TYPE "UDT1800_FLT_Machine"
VERSION : 0.1
   STRUCT
      Data_lost_after_erasing : Bool;   // Data_lost_after_erasing S7-CPU (1)
      Fuse_broken : Bool;   // Fuse broken machine (3)
      Connection_To_PC_lost : Bool;   // Connection to PC lost (3)
      Door_Swichtcabinet_open : Bool;   // Door swichtcabinet open(3)
      Air_dryer : Bool;   // Air dryer (3)
      Controlvoltage : Bool;   // Controlvoltage missing (M)
      CylinderServiceNotPermit : Bool;   // Operationmode cylinder service not permitted (1)
      Fuse_brocken_Mixinghead : Bool;   // Fuse broken mixinghead (3)
      Heating : Bool;   // Heating of machine overload (3)
      SGM_Faulty : Bool;   // Extrusion machine faulty (3)
      F_CoolingDevice : Bool;   // Compressor cooling device (3)
      WrongMH_No : Bool;   // Wrong mixinghead number (1)
      PlasmaFaulty : Bool;   // Plasma unit faulty (3)
      DrainingTank : Bool;   // Draining of a tank selected (M)
      SGM_AutomatcMissing : Bool;   // Extrusion machine not in automatic maode (3)
      Spare_1_7 : Bool;
      EmergencyStop : Struct   // Emergency stop general (M)
         Machine : Bool;   // Emergency stop nachine
         Switch_Cabinet : Bool;   // Emergency stop switch cabinet
         Operation_Panel : Bool;   // Emergency stop operation panel
         Monitor_2 : Bool;   // Emergency stop monitor_2
         Tank : Bool;   // Emergency stop tank
         MH_Cleaner_1 : Bool;   // Emergency stop mixinghead cleaner 1
         MH_Cleaner_2 : Bool;   // Emergency stop mixinghead cleaner 2
         Roboter_1 : Bool;   // Emergency stop Robot 1
         Roboter_2 : Bool;   // Emergency stop Robot 2
         ContStation_C1 : Bool;   // Emergency stop container station component 1
         ContStation_C2 : Bool;   // Emergency stop container station component 2
         External_Plant_1 : Bool;   // Emergency stop external plant 1
         External_Plant_2 : Bool;   // Emergency stop external plant 2
         ColorUnit_01 : Bool;   // Emergency stop color unit 1
         ColorUnit_02 : Bool;   // Emergency stop color unit 2
         AdditionalComponent : Bool;   // Emergency stop additional component
      END_STRUCT;
      OpMode_Test : Bool;   // Operation mode test is selected (M)
      Weekend_Mode : Bool;   // Weekende mode is active (M)
      Interface_PC : Bool;
      BufferBattery : Bool;
      AutoStop : Bool;   // AutoStop active (M)
      FLT_pre_alarm_pentan : Bool;   // Fault pre alarm pentan (3)
      FLT_alarm_pentan : Bool;   // Fault alarm pentan (1)
      P_AirSupply : Bool;   // Fault supply air pressure too low (3)
      FaultPC_Level_1 : Bool;
      FaultPC_Level_2 : Bool;
      FaultPC_Level_3 : Bool;
      Spare_13_3 : Bool;
      BufferShotDataFull : Bool;
      TransferFaultMMC : Bool;
      Fault_Watchdog : Bool;
      RefillStationNotReady : Bool;
      ShotTimeTooShort : Bool;
      CantDeleteTool : Bool;
      Pneumatik_1 : Bool;
      Pneumatik_2 : Bool;
      Spare_14_04 : Bool;
      Spare_14_05 : Bool;
      Spare_14_06 : Bool;
      Spare_14_07 : Bool;
      TimeValueIntervallNOK : Bool;
      Spare_15_01 : Bool;
      Spare_15_02 : Bool;
      Spare_15_03 : Bool;
      Spare_15_04 : Bool;
      Spare_15_05 : Bool;
      Spare_15_06 : Bool;
      Spare_15_07 : Bool;
      Spare_16_00 : Bool;
      Spare_16_01 : Bool;
      Spare_16_02 : Bool;
      Spare_16_03 : Bool;
      Spare_16_04 : Bool;
      Spare_16_05 : Bool;
      Spare_16_06 : Bool;
      Spare_16_07 : Bool;
      Spare_17_00 : Bool;
      Spare_17_01 : Bool;
      Spare_17_02 : Bool;
      Spare_17_03 : Bool;
      Spare_17_04 : Bool;
      Spare_17_05 : Bool;
      Spare_17_06 : Bool;
      Spare_17_07 : Bool;
   END_STRUCT;
END_TYPE

TYPE "UDT1801_FLT_auxDrive"
VERSION : 0.1
   STRUCT
      FLT_Motorprotection : Bool;   // Fault motorprotection
      FLT_FrequencyConverter : Bool;   // Fault frequency converter
      FLT_MaxP_MaxLTripTray : Bool;   // Max. level trip tray or max. pressure component
      FLT_Dryrunsafety : Bool;   // Fault dryrun safety
      FLT_wrong_Timevalue : Bool;   // Wrong timevalue at run- and pause time (3)
      FLT_MaxPressureDiff : Bool;   // Fault: Max. pressure difference at filter
      Mes_Min_temp : Bool;   // Message min. temperature not reached to start drive
      FLT_MotorFan : Bool;   // Fault: Motorprotection external fan of motor
      Mes_Min_Level : Bool;   // Message min. level not reached to start drive
      FLT_No_Barrel : Bool;   // Fault: No barrel existing during filling request
      Mes_No_Barrel : Bool;   // Message: No barrel existing
      Spare_1_3 : Bool;
      Spare_1_4 : Bool;
      Spare_1_5 : Bool;
      Spare_1_6 : Bool;
      Spare_1_7 : Bool;
   END_STRUCT;
END_TYPE

TYPE "UDT1802_FLT_Tank_Refill"
VERSION : 0.1
   STRUCT
      FLT_Min_Level : Bool;   // Filling level tank below minimum (1)
      FLT_Max_Level : Bool;   // Filling level tank over maximum (3)
      FLT_Fillingtime_to_long : Bool;   // Maximum fillingtime exceeded (3)
      FLT_Max_Level_Triptray : Bool;   // Maximum level triptray (3)
      FLT_Min_Level_Cycle : Bool;   // Level tank below minimum during foaming cycle (2)
      FLT_Max_Level_Pistonm : Bool;   // Max level tank at piston machine (1)
      FLT_Max_Level_Tt_Pistonm : Bool;   // Maximum level triptray at piston machine (2)
      FLT_LevelSensor_broken_wire : Bool;   // There is no connection to the level sensor (3)
      FLT_Filling_Valve_AS : Bool;   // Fault position filling valve (3)
      FLT_PreWarning_Min_Level : Bool;   // Pre Warning min. level reached (3)
      FLT_Spare_11 : Bool;
      FLT_Spare_12 : Bool;
      FLT_Spare_13 : Bool;
      FLT_supply_nucleation : Bool;   // Fault supply nucleation (3)
      FLT_NucleationSensor_broken_wire : Bool;   // There is no connection to the nucleation sensor (3)
      FLT_nucleation : Bool;   // Fault Message from nucleation (3)
   END_STRUCT;
END_TYPE

TYPE "UDT1803_FLT_RefilStation"
VERSION : 0.1
   STRUCT
      Message_No_drum : Bool;   // Meldung: Es ist kein Faß in der Containerstation vorhanden
      Message_Spare : Bool;
      FLT_Min_Pressure_Air : Bool;   // Störung: Eingestellter min. Druck der Luftversorgung unterschritten (3)
      FLT_MinPressureAirPump : Bool;
      FLT_Heat1 : Bool;
      FLT_Heat2 : Bool;
      FLT_Spare06 : Bool;
      FLT_Spare07 : Bool;
      FLT_Spare10 : Bool;
      FLT_Drum_is_empty : Bool;   // Störung: Das Faß in der Containerstatiuon ist leer! Bitte wechseln! (3)
      FLT_Dryprotection_RCP : Bool;   // Störung: Der Trockenlaufschutz an der Kreislaufpumpe hat angesprochen (3)
      FLT_MaxPressureComponent : Bool;   // Störung: Der Komponentendruck in der Kreislaufleitung wurde überschritten (3)
      EmergencyStop : Bool;
      FLT_Spare_1_5 : Bool;
      FLT_Spare_1_6 : Bool;
      FLT_Spare_1_7 : Bool;
      Agitator : "UDT1801_FLT_auxDrive";
      Pump : "UDT1801_FLT_auxDrive";
      Filling : "UDT1802_FLT_Tank_Refill";
   END_STRUCT;
END_TYPE

TYPE "UDT1804_FLT_Controller"
VERSION : 0.1
   STRUCT
      Sensor_FLT_broken_wire : Bool;   // There is no connection to the sensor (3)
      Warning_limit_plus : Bool;   // The lower warning limit of the processvalue under run (3)
      Warning_limit_minus : Bool;   // The upper warning limit of the processvalue is exceeded (3)
      Alarm_limit_plus : Bool;   // The lower alarm limit of the processvalue under run(1)
      Alarm_limit_minus : Bool;   // The upper alarm limit of the processvalue is exceeded (1)
      Controller_at_limit : Bool;   // Controller at limit (3)
      spare06 : Bool;
      Fuse_TemperingUnit : Bool;   // Fault Tempering Unit (3)
      Fuse_TemperingOverLoad : Bool;   // Overload tempering unit (3)
      lower_limit : Bool;   // controler value under limit (3)
      upper_limit : Bool;   // controler value over limit (3)
      HW_Limit : Bool;   // Controller at hardware limit (3)
      NoSetValue : Bool;   // Set value = 0! No function (3)
      spare013 : Bool;
      spare014 : Bool;
      spare015 : Bool;
   END_STRUCT;
END_TYPE

TYPE "UDT1805_FLT_PB_DP"
VERSION : 0.1
   STRUCT
      Member : Array[1..128] of Bool;
   END_STRUCT;
END_TYPE

TYPE "UDT1806_FLT_Vacuum"
VERSION : 0.1
   STRUCT
      FLT_PVacuum : Bool;
      Motorprotection : Bool;
      Spare2 : Bool;
      Spare3 : Bool;
      Spare4 : Bool;
      Spare5 : Bool;
      Spare6 : Bool;
      Spare7 : Bool;
   END_STRUCT;
END_TYPE

TYPE "UDT1807_FaultMicroMeter"
VERSION : 0.1
   STRUCT
      MultibleAllocation : Bool;   // Allocation of metering unit at mixing head more then one connector (1)
      NotSelected : Bool;   // Selection of metering unit by switch missing
      PowerSupply : Bool;   // Power supply metering unit faulty (1)
      Watchdog : Bool;   // No sign of live signal from metering unit
      NotOperative : Bool;   // Metering unit not ready for operation (1)
      NotAllocated : Bool;   // Metering unit not allocated to mixinghead connector (1)
      Spare01 : Bool;
      Spare02 : Bool;
      Spare10 : Bool;
      Spare11 : Bool;
      Spare12 : Bool;
      Spare13 : Bool;
      Spare14 : Bool;
      Spare15 : Bool;
      Spare16 : Bool;
      Spare17 : Bool;
   END_STRUCT;
END_TYPE

TYPE "UDT1801_Agitator"
VERSION : 0.1
   STRUCT
      FLT_Motorprotection : Bool;   // Fault motorprotection
      FLT_FrequencyConverter : Bool;   // Fault frequency converter
      FLT_MaxLTripTray : Bool;   // Max. level trip tray
      FLT_wrong_Timevalue : Bool;   // Wrong timevalue at run- and pause time (3)
      FLT_MaxPressureDiff : Bool;   // Fault: Max. pressure difference at filter
      Mes_Min_temp : Bool;   // Message min. temperature not reached to start drive
      FLT_MotorFan : Bool;   // Fault: Motorprotection external fan of motor
      Mes_Min_Level : Bool;   // Message min. level not reached to start drive
      Mes_Min_Temp_1 : Bool;   // Message min. temperature not reached
      Spare_1_2 : Bool;
      Spare_1_3 : Bool;
      Spare_1_4 : Bool;
      Spare_1_5 : Bool;
      Spare_1_6 : Bool;
      Spare_1_7 : Bool;
   END_STRUCT;
END_TYPE

TYPE "UDT1809_FLT_CoverLift"
VERSION : 0.1
   STRUCT
      RunTimeCoverLifting : Bool;
      RunTimeCoverDropping : Bool;
      PressureAirCoverLift : Bool;
      Spare03 : Bool;
      Spare04 : Bool;
      Spare05 : Bool;
      Spare06 : Bool;
      Spare07 : Bool;
   END_STRUCT;
END_TYPE

TYPE "UDT1801_EdgeFilter"
VERSION : 0.1
   STRUCT
      FLT_Motorprotection : Bool;   // Fault motorprotection
      FLT_MaxPressureDiff : Bool;   // Fault: Max. pressure difference at filter
      FLT_wrong_Timevalue : Bool;   // Wrong timevalue at run- and pause time (3)
      Spare_1_3 : Bool;
      Spare_1_4 : Bool;
      Spare_1_5 : Bool;
      Spare_1_6 : Bool;
      Spare_1_7 : Bool;
   END_STRUCT;
END_TYPE

TYPE "UDT1811_GenAuxDrives"
VERSION : 0.1
   STRUCT
      FanHousing : "UDT1801_FLT_auxDrive";
      AuxDrive_Spare01 : "UDT1801_FLT_auxDrive";
      AuxDrive_Spare02 : "UDT1801_FLT_auxDrive";
      AuxDrive_Spare03 : "UDT1801_FLT_auxDrive";
      AuxDrive_Spare04 : "UDT1801_FLT_auxDrive";
      AuxDrive_Spare05 : "UDT1801_FLT_auxDrive";
      AuxDrive_Spare06 : "UDT1801_FLT_auxDrive";
      AuxDrive_Spare07 : "UDT1801_FLT_auxDrive";
      AuxDrive_Spare08 : "UDT1801_FLT_auxDrive";
      AuxDrive_Spare09 : "UDT1801_FLT_auxDrive";
      AuxDrive_Spare10 : "UDT1801_FLT_auxDrive";
   END_STRUCT;
END_TYPE

TYPE "UDT1801_FeedingPump"
VERSION : 0.1
   STRUCT
      FLT_Motorprotection : Bool;   // Fault motorprotection
      FLT_FrequencyConverter : Bool;   // Fault frequency converter
      FLT_MaxLTripTray : Bool;   // Max. level trip tray
      FLT_Dryrunsafety : Bool;   // Fault dryrun safety
      FLT_wrong_Timevalue : Bool;   // Wrong timevalue at run- and pause time (3)
      FLT_MaxPressure : Bool;   // Max. pressure component
      Mes_Min_temp : Bool;   // Message min. temperature not reached to start drive
      FLT_MotorFan : Bool;   // Fault: Motorprotection external fan of motor
      Spare_09 : Bool;
      Spare_10 : Bool;
      Spare_11 : Bool;
      Spare_12 : Bool;
      Spare_13 : Bool;
      Spare_14 : Bool;
      Spare_15 : Bool;
      Spare_16 : Bool;
   END_STRUCT;
END_TYPE

TYPE "Fanuc_Faults"
VERSION : 0.1
   STRUCT
      doSysError : Bool;
      No_Cycle_Program : Bool;
      Program_transmission : Bool;
      No_Moulds_Faulty : Bool;
      No_ShotTimes_Faulty : Bool;
      ShotTime_Faulty : Bool;
      MouldSelection_Faulty : Bool;
      Roboter_Stopped : Bool;
      FLT_System : Bool;
      FLT_Interface : Bool;
      FLT_Fuse_Supply : Bool;
      FLT_doAction_01 : Bool;
      FLT_RobnotHP_Cyclestart : Bool;   // Roboter not in home position at cycle start
      FLT_Rob_not_ready_for_PU : Bool;   // Roboter not ready
      FLT_OldProgsNotReady : Bool;   // New programs for robot detected, while old programs still active (1)
      FLT_PUnotReadyForShot : Bool;   // robot starts next shot but PU is not ready yet (1)
      FLT_RobStoppedInProd : Bool;   // Robot stopped while production is runnung (1)
      FLT_TPOnInProd : Bool;   // Teach pendant is on in production (1)
      FLT_PrgNotExisting : Bool;   // A requested program is not existing in the robot (1)
      FLT_RobInClosingMould : Bool;   // The robot is still in a mould that is about to close (Worldzone) (1)
      FLT_RobInClosingTrolley : Bool;   // The trolley number the robot reports back is in closing area (1)
      FLT_Stepnumber_not_zero : Bool;   // Stepnumber of step control not zero
      Roboter_not_in_automatic : Bool;
      RobotProgramNotRunning : Bool;
      FaultNumber : Byte;
   END_STRUCT;
END_TYPE

TYPE "UDT1816_FLT_IF_SP_MC"
VERSION : 0.1
   STRUCT
      Fault_IF : Bool;   // Fault as interface was at first position (3)
      FLT_pouring_release : Bool;   // Foaming release was set to zero (3)
      FLT_SWU_release : Bool;   // SWU release was set to zero. (3)
      FLT_Stop_while_selected : Bool;   // Stop button was set to zero (3)
      FLT_op_mode_O : Bool;   // Key switch manual/automatic was set to zero (3)
      FLT_Cycle_release : Bool;   // Release foaming cycle was set to zero (3)
      FLT_Communication : Bool;   // Fault communication mc (3)
      FLT_NoCupAtTestshotposition : Bool;   // Fault that there is no cup at the testshot position
      Spare_1_0 : Bool;
      Spare_1_1 : Bool;
      Spare_1_2 : Bool;
      Spare_1_3 : Bool;
      Spare_1_4 : Bool;
      Spare_1_5 : Bool;
      Spare_1_6 : Bool;
      Spare_1_7 : Bool;
   END_STRUCT;
END_TYPE

TYPE "UDT1817_FLT_IF_extPlant"
VERSION : 0.1
   STRUCT
      FLT_Strobe : Bool;   // The signal strobe appears before the plant is ready to operate (3)
      FLT_Strobe_inv : Bool;   // The signal strobe inverse appears before the plant is ready to operate (3)
      MSG_AP_not_OK : Bool;   // The external plant not at automatic mode // Message
      FLT_AP_not_OK : Bool;   // The external plant is not at automatic mode during release of cycle // (3)
      FLT_no_number : Bool;   // Strobe set but there is no or a wrong program number (3)
      FLT_inverse_number : Bool;   // The inverse program number was wrong (3)
      FLT_Parity_Bit : Bool;   // Parity bit was wrong (3)
      FLT_Start_Shot : Bool;   // Signal start shot is set at the start of foaming cycle (3)
      FLT_Cycle_Stoped : Bool;   // A registerd interface will be taken off the liste (3)
      FLT_Watchdog : Bool;   // check watchdog signal from the external plant
      Reserve2 : Bool;
      Reserve3 : Bool;
      Reserve4 : Bool;
      Reserve5 : Bool;
      Reserve6 : Bool;
      Reserve7 : Bool;
   END_STRUCT;
END_TYPE

TYPE "UDT1818_FLT_RinsingStat"
VERSION : 0.1
   STRUCT
      Warning_Min_Level : Bool;   // Warning: Level tank below min. value
      FLT_Min_Level : Bool;   // Fault: Min. level tank below (> 5 min.)
      Warning_Min_Temp : Bool;   // Warning: Temperatur tank below min. value
      FLT_Min_Temp : Bool;   // Fault: Min. temperatur tank below (> 5 min.)
      FLT_Min_Pressure : Bool;   // Fault: Min. cleaning pressure not reached
      FLT_Max_Pressure : Bool;   // Fault: Maximum cleaning pressure reached
      FLT_SystemPressure : Bool;   // Fault: Min. pressure air wurde unterschritten
      FLT_TimeValue_Null : Bool;   // Fault: Timevalue of MH (spray) = 0
      FLT_RinsingPump : Bool;   // Fault: motorprotection resing pump
      Spare_11 : Bool;   // --------------
      Spare_12 : Bool;   // --------------
      Spare_13 : Bool;   // --------------
      Spare_14 : Bool;   // --------------
      Spare_15 : Bool;   // --------------
      Spare_16 : Bool;   // --------------
      Spare_17 : Bool;   // --------------
   END_STRUCT;
END_TYPE

TYPE "UDT1819_FLT_PouringCycle"
VERSION : 0.1
   STRUCT
      FLT_KLZ_0 : Bool;   // Fault no valid time value (3)
      FLT_Max_Waittime : Bool;   // Fault maximum waiting time after CLT1 or CLT3 exceeded (3)
      FLT_Max_Shottime : Bool;   // Fault actual foamingtime exceeded limit (1)
      FLT_OP_Mode : Bool;   // Fault operation mode changed during foaming cycle (1)
      Reserve1 : Bool;
      Reserve2 : Bool;
      Reserve3 : Bool;
      FLT_CompAllocation : Bool;   // Pumpno. or tankno. allocated = 0
      FLT_NewNoTooEarly : Bool;   // New station number detected while old number still active
      FLT_WRongStationNumber : Bool;   // Wrong station no or mistake in station list
      FLT_WrongToolNumber : Bool;   // Wrong tool no or mistake in tool list
      FLT_WrongShotNumber : Bool;   // Wrong shot number in tool data
      FLT_WrongMixingheadNumber : Bool;   // Wrong mixinghead number at tool data
      FLT_TransferShotResult : Bool;   // Fault transfer shot result from buffer to PUC-DB
      FLT_BufferShotResultFull : Bool;
      Spare_1_7 : Bool;
   END_STRUCT;
END_TYPE

TYPE "UDT1820_FLT_ProcessValue"
VERSION : 0.1
   STRUCT
      Sensor_FLT_broken_wire : Bool;   // There is no connection to the sensor (3)
      Warning_limit_plus : Bool;   // The lower warning limit of the processvalue under run (3)
      Warning_limit_minus : Bool;   // The upper warning limit of the processvalue is exceeded (3)
      Alarm_limit_plus : Bool;   // The lower alarm limit of the processvalue under run(1)
      Alarm_limit_minus : Bool;   // The upper alarm limit of the processvalue is exceeded (1)
      Controller_at_limit : Bool;   // Controller at limit (3)
      Spare_0_6 : Bool;
      Fuse_TemperingOverLoad : Bool;   // Overload tempering unit (3)
      Spare_1_0 : Bool;
      Spare_1_1 : Bool;
      Spare_1_2 : Bool;
      Spare_1_3 : Bool;
      Spare_1_4 : Bool;
      Spare_1_5 : Bool;
      Spare_1_6 : Bool;
      Spare_1_7 : Bool;
   END_STRUCT;
END_TYPE

TYPE "UDT1821_FLT_MH_Hydraulic"
VERSION : 0.1
   STRUCT
      FLT_Motorprotection : Bool;   // Fault motor protection hydraulic (1)
      FLT_Min_Level : Bool;   // Fault min level oil tank hydraulic (1)
      FLT_WRN_C_Max : Bool;   // Fault warning temperature hydraulic oil (2)
      FLT_C_Max : Bool;   // Fault temperature hydraulic oil more than 5 min.too high (1)
      FLT_Filter_HP : Bool;   // Fault pre run high pressure filter hydraulic soild (3)
      FLT_Filter_backflow : Bool;   // Fault back flow filter hydraulic soild (3)
      FLT_cable_break : Bool;   // Fault cable break pressure switch (1)
      FLT_P_Max : Bool;   // Fault maximum pressure hydraulic not reached (1)
      FLT_Moog_Filter : Bool;   // Fault moog filter hydraulic (3)
      FLT_MotorProtFilterPump : Bool;   // Fault motor protection filter pump (1)
      FLT_MinLevelFilterPump : Bool;   // Fault minimum level on side of filter pump (1)
      FLT_MaxLevelFilterPump : Bool;   // Fault maximum level on side of filter pump (1)
      FLT_FilterBypass : Bool;   // Fault filter bypass soild (3)
      Spare14 : Bool;
      Spare15 : Bool;
      Spare16 : Bool;
   END_STRUCT;
END_TYPE

TYPE "UDT1822_FLT_PV_Flow"
VERSION : 0.1
   STRUCT
      Sensor_FLT_broken_wire : Bool;   // Wire break Sensor (3)
      Warning_limit_plus : Bool;   // Warning limit exceeded (3)
      Warning_limit_minus : Bool;   // Warning limit underflowed (3)
      Alarm_limit_plus : Bool;   // Alarm limit exceeded (1)
      Alarm_limit_minus : Bool;   // Alarm limit underflowed (1)
      Controller_at_limit : Bool;   // Flow controler at the limit (3)
      Reserve1 : Bool;
      Reserve2 : Bool;
      Spare_1_0 : Bool;
      Warning_limit_plus_MR : Bool;   // Warning limit exceeded mixing ratio (3)
      Warning_limit_minus_MR : Bool;   // Warning limit underflow mixing ratio (3)
      Alarm_limit_plus_MR : Bool;   // Alarm limit exceeded mixing ratio (1)
      Alarm_limit_minus_MR : Bool;   // Alarm limit underflow mixing ratio (1)
      Spare_1_5 : Bool;
      Spare_1_6 : Bool;
      Spare_1_7 : Bool;
   END_STRUCT;
END_TYPE

TYPE "UDT1823_FLT_Chain"
VERSION : 0.1
   STRUCT
      FLT_pressure : Bool;   // Pressure switch does not work correctly (1)
      FLT_mot_prot : Bool;   // Motor protection (1)
      FLT_min_level : Bool;   // Min level oil (1)
      FLT_filter : Bool;   // Filter contaminated (3)
      FLT_C_Max : Bool;   // Fault max temperature (1)
      WRN_C_Max : Bool;   // Warning max temperature (2)
      FLT_chain_too_long : Bool;   // Chain too long (1)
      Spare0_7 : Bool;
      FLT_ConveyorPosition : Bool;   // Fault with detection of conveyor position (1)
      MSG_ConvPosUnKnown : Bool;   // Message: position of conveyor is unknown (4)
      Spare1_2 : Bool;
      FLT_PowerRail : Bool;   // Motor protection power rail of conveyor (1)
      Spare1_4 : Bool;
      Spare1_5 : Bool;
      FLT_MinLevelLubrication : Bool;   // Min level of chain lubrication (3)
      FLT_NoPulsesLubrication : Bool;   // No pulses to start chain lubrication (3)
   END_STRUCT;
END_TYPE

TYPE "UDT1824_FLT_GBE"
VERSION : 0.1
   STRUCT
      EmergencyStop : Bool;   // Emergency Stop from GBE
      FLT_Supply : Bool;   // Fault Supply from GBE
      FLT_Interface : Bool;   // Fault from Interface GBE
      Spare_0_3 : Bool;
      Spare_0_4 : Bool;
      Spare_0_5 : Bool;
      Spare_0_6 : Bool;
      Spare_0_7 : Bool;
      Spare_1_0 : Bool;
      Spare_1_1 : Bool;
      Spare_1_2 : Bool;
      Spare_1_3 : Bool;
      Spare_1_4 : Bool;
      Spare_1_5 : Bool;
      Spare_1_6 : Bool;
      Spare_1_7 : Bool;
   END_STRUCT;
END_TYPE

TYPE "UDT1826_FLT_LeakageMonit"
VERSION : 0.1
   STRUCT
      Fault_Leakage : Bool;
      Fault_Threshold : Bool;
      Spare_02 : Bool;
      Spare_03 : Bool;
      Spare_04 : Bool;
      Spare_05 : Bool;
      Spare_06 : Bool;
      Spare_07 : Bool;
      Spare_010 : Bool;
      Spare_011 : Bool;
      Spare_012 : Bool;
      Spare_013 : Bool;
      Spare_014 : Bool;
      Spare_015 : Bool;
      Spare_016 : Bool;
      Spare_017 : Bool;
   END_STRUCT;
END_TYPE

TYPE "UDT1827_ErrorMovMouldMC"
VERSION : 0.1
   STRUCT
      ErrorStateToolBin : Struct
         MC_Motion_01_OP : Bool;   // 01: Lid closed
         MC_Motion_02_OP : Bool;   // 02: Left lock closed
         MC_Motion_03_OP : Bool;   // 03: Right lock closed
         MC_Motion_04_OP : Bool;   // 04: Left air cushion inflated
         MC_Motion_05_OP : Bool;   // 05: Right air cushion inflated
         MC_Motion_06_OP : Bool;   // 06:
         MC_Motion_07_OP : Bool;   // 07:
         MC_Motion_08_OP : Bool;   // 08:
         MC_Motion_09_OP : Bool;   // 09:
         MC_Motion_10_OP : Bool;   // 10:
         MC_Motion_11_OP : Bool;   // 11:
         MC_Motion_12_OP : Bool;   // 12:
         MC_Motion_13_OP : Bool;   // 13:
         MC_Motion_14_OP : Bool;   // 14: Mould existing left side
         MC_Motion_15_OP : Bool;   // 15: Mould existing right side
         MC_Motion_16_OP : Bool;   // 16: Cassette existing
         MC_Motion_01_BP : Bool;   // 17: Lid opened
         MC_Motion_02_BP : Bool;   // 18: Left lock opened
         MC_Motion_03_BP : Bool;   // 19: Right lock opened
         MC_Motion_04_BP : Bool;   // 20: Left air cushion bleeded
         MC_Motion_05_BP : Bool;   // 21: Right air cushion bleeded
         MC_Motion_06_BP : Bool;   // 22:
         MC_Motion_07_BP : Bool;   // 23:
         MC_Motion_08_BP : Bool;   // 24:
         MC_Motion_09_BP : Bool;   // 25:
         MC_Motion_10_BP : Bool;   // 26:
         MC_Motion_11_BP : Bool;   // 27:
         MC_Motion_12_BP : Bool;   // 28:
         MC_Motion_13_BP : Bool;   // 29:
         MC_Motion_14_BP : Bool;   // 30:
         MC_Motion_15_BP : Bool;   // 31:
         MC_Motion_16_BP : Bool;   // 32:
         Mould_Motion_01_OP : Bool;   // 33: 3rd part of tool in
         Mould_Motion_02_OP : Bool;   // 34: Autovent in
         Mould_Motion_03_OP : Bool;   // 35:
         Mould_Motion_04_OP : Bool;   // 36:
         Mould_Motion_05_OP : Bool;   // 37:
         Mould_Motion_06_OP : Bool;   // 38:
         Mould_Motion_07_OP : Bool;   // 39:
         Mould_Motion_08_OP : Bool;   // 40:
         Mould_Motion_09_OP : Bool;   // 41:
         Mould_Motion_10_OP : Bool;   // 42:
         Mould_Motion_11_OP : Bool;   // 43:
         Mould_Motion_12_OP : Bool;   // 44:
         Mould_Motion_13_OP : Bool;   // 45:
         Mould_Motion_14_OP : Bool;   // 46:
         Mould_Motion_15_OP : Bool;   // 47:
         Mould_Motion_16_OP : Bool;   // 48:
         Mould_Motion_01_BP : Bool;   // 49: 3rd part of tool out
         Mould_Motion_02_BP : Bool;   // 50: Autovent out
         Mould_Motion_03_BP : Bool;   // 51:
         Mould_Motion_04_BP : Bool;   // 52:
         Mould_Motion_05_BP : Bool;   // 53:
         Mould_Motion_06_BP : Bool;   // 54:
         Mould_Motion_07_BP : Bool;   // 55:
         Mould_Motion_08_BP : Bool;   // 56:
         Mould_Motion_09_BP : Bool;   // 57:
         Mould_Motion_10_BP : Bool;   // 58:
         Mould_Motion_11_BP : Bool;   // 59:
         Mould_Motion_12_BP : Bool;   // 60:
         Mould_Motion_13_BP : Bool;   // 61:
         Mould_Motion_14_BP : Bool;   // 62:
         Mould_Motion_15_BP : Bool;   // 63:
         Mould_Motion_16_BP : Bool;   // 64:
         GeneralStatus01 : Bool;   // 65: Foam is in the mould
         GeneralStatus02 : Bool;   // 66: Part was taken out of the mould
         GeneralStatus03 : Bool;   // 67: The waiting time for venting is active
         GeneralStatus04 : Bool;   // 68: Venting stroke is active
         GeneralStatus05 : Bool;   // 69: Reaction time is running
         GeneralStatus06 : Bool;   // 70:
         GeneralStatus07 : Bool;   // 71:
         GeneralStatus08 : Bool;   // 72:
         GeneralStatus09 : Bool;   // 73:
         GeneralStatus10 : Bool;   // 74:
         GeneralStatus11 : Bool;   // 75:
         GeneralStatus12 : Bool;   // 76:
         GeneralStatus13 : Bool;   // 77:
         GeneralStatus14 : Bool;   // 78:
         GeneralStatus15 : Bool;   // 79: Mould is not in handling area (1 safety switch per trolley)
         GeneralStatus16 : Bool;   // 80:
         Parity_Mouldcoding : Bool;   // Störung Parität Formcodierung [1]
         Transmission_Mouldcoding : Bool;   // Fehler beim Senden der Codierung an PU [1]
         NoMouldcodingHigh : Bool;   // Formcodierung zu groß [1]
         MouldcodingMissing : Bool;   // Formcodierung fehlt [1]
         AllocationMH_Mould : Bool;   // Die Anwahl der Mischköpfe und der Formen stimmt nicht überein [1]
         FuseTemperingUnit : Bool;   // Sicherung Temperiergerät [3]
         Spare10_6 : Bool;
         Spare10_7 : Bool;
         Spare11_0 : Bool;
         Spare11_1 : Bool;
         Spare11_2 : Bool;
         Spare11_3 : Bool;
         Spare11_4 : Bool;
         Spare11_5 : Bool;
         Spare11_6 : Bool;
         Spare11_7 : Bool;
      END_STRUCT;
   END_STRUCT;
END_TYPE

TYPE "UDT1828_ErrorMC"
VERSION : 0.1
   STRUCT
      MotorprotectionVacuum : Bool;
      PressureBuildUpVacuum : Bool;
      RestartDelayVacuum : Bool;
      FoamingMachineNotOK : Bool;
      FuseGeneral : Bool;
      FuseTemperingUnit : Bool;
      LightSwitchNotAckn : Bool;
      SaftyDoorMCNotAckn01 : Bool;
      SaftyDoorMCNotAckn02 : Bool;
      EmergenStopSwitchCabinet : Bool;
      EmergenStopHydraulic : Bool;
      EmergenStopOpanel : Bool;
      LiftGateNotClosed01 : Bool;
      LiftGateNotClosed02 : Bool;
      Flap01 : Bool;   // Pendelklappe
      Flap02 : Bool;   // Pendelklappe
      UpperLimitFlow : Bool;   // Upper limit discharge flow of all components
      LowerLimitFlow : Bool;   // Lower limit discharge flow of all components
      NoPressureSensorSelected : Bool;
      Spare23 : Bool;
      Spare24 : Bool;
      Spare25 : Bool;
      Spare26 : Bool;
      Spare27 : Bool;
      Spare30 : Bool;
      Spare31 : Bool;
      Spare32 : Bool;
      Spare33 : Bool;
      Spare34 : Bool;
      Spare35 : Bool;
      Spare36 : Bool;
      Spare37 : Bool;
   END_STRUCT;
END_TYPE

TYPE "UDT1829_ErrorDriveConv"
VERSION : 0.1
   STRUCT
      FLT_FreqConverter : Bool;   // Frequency converter not ready for operation (1)
      FLT_Motor : Bool;   // Motor protection (1)
      FLT_Fan : Bool;   // Fault external fan of Motor (2)
      Spare0_3 : Bool;
      Spare0_4 : Bool;
      FLT_FromIPos : Bool;   // Error message from frequency converter (1)
      FLT_PosCheckIni : Bool;   // Proximity switch for position check is not on (1)
      FLT_PosCheckIniAllwaysOn : Bool;   // Proximity switch for position check is allways on (1)
      Spare1_0 : Bool;
      Spare1_1 : Bool;
      Spare1_2 : Bool;
      Spare1_3 : Bool;
      Spare1_4 : Bool;
      Spare1_5 : Bool;
      Spare1_6 : Bool;
      Spare1_7 : Bool;
   END_STRUCT;
END_TYPE

TYPE "UDT1830_FLT_PipesHeating"
VERSION : 0.1
   STRUCT
      Pipe01 : "UDT1820_FLT_ProcessValue";
      Pipe02 : "UDT1820_FLT_ProcessValue";
   END_STRUCT;
END_TYPE

TYPE "UDT1831_FLT_EPS_Robot"
VERSION : 0.1
   STRUCT
      FLT_SyncSwitch : Bool;   // [3] EPS Sync Switch damaged or Snyc Position robot not ok
      FLT_NotSynchonized : Bool;   // [3] EPS is not synchronized
      FLT_RestartRequired : Bool;   // [3] EPS demanded Restart (Warmstart)
      FLT_PreWarnIsAktiv : Bool;   // [4] EPS is only a short time synchronized
      FLT_CollisionProtection : Bool;   // [4] Collision protection as triggered // Rammschutz
      Spare_0_5 : Bool;
      Spare_0_6 : Bool;
      Spare_0_7 : Bool;
      FHM_FLT_SyncSwitch : Bool;
      FHM_FLT_NotSynchonized : Bool;
      FHM_FLT_RestartRequired : Bool;
      FHM_FLT_PreWarnIsAktiv : Bool;
      FHM_FLT_CollisionProtect : Bool;
      FHM_Spare_1_5 : Bool;
      FHM_Spare_1_6 : Bool;
      FHM_Spare_1_7 : Bool;
   END_STRUCT;
END_TYPE

TYPE "UDT1841_FLT_SWU"
VERSION : 0.1
   STRUCT
      FLT_open_SWU_disabelt : Bool;   // Fault selected switch over unit disabelt (1)
      FLT_No_SWU_selected : Bool;   // Fault no switch over unit selected (1)
      FLT_Sel_SWU_not_released : Bool;   // Fault selected switch over unit not released (1)
      spare_0_3 : Bool;
      spare_0_4 : Bool;
      spare_0_5 : Bool;
      spare_0_6 : Bool;
      spare_0_7 : Bool;
      spare_1_0 : Bool;
      spare_1_1 : Bool;
      spare_1_2 : Bool;
      spare_1_3 : Bool;
      spare_1_4 : Bool;
      spare_1_5 : Bool;
      spare_1_6 : Bool;
      spare_1_7 : Bool;
   END_STRUCT;
END_TYPE

TYPE "UDT1842_FLT_MH_Control"
VERSION : 0.1
   STRUCT
      FLT_MH_dontOpen : Bool;   // Mixinghead do not open (1)
      FLT_MH_dontClose : Bool;   // Mixinghead do not close (1)
      FLT_ShotStopped : Bool;   // Break during shot (3)
      FLT_MH_OpenWOactivation : Bool;   // Mixinghead open with out activation (1)
      FLT_MH_CloseDuringShot : Bool;   // Mixinghead close during shot (3)
      WRN_ShotTimeShort : Bool;   // Warning shot time too short (3)
      WRN_ShotTimeLong : Bool;   // Warning shot time too long (3)
      FLT_ShotTimeShort : Bool;   // Fault shot time too short (3)
      FLT_MH_bounce : Bool;   // MH bounce during opening or closing (3)
      FLT_RT_Lock : Bool;   // Time locking mixinghead takes too long (1)
      FLT_RT_Unlock : Bool;   // Time unlocking mixinghead takes too long (1)
      WRN_NozzleLeakageTest_active : Bool;   // The nozzle leakage test is active. Nozzles and bypasses are closed
      Spare_1_4 : Bool;
      Spare_1_5 : Bool;
      Spare_1_6 : Bool;
      FLTCompNotOnThisMH : Bool;   // Component in shot is not connected to this mixinghead
   END_STRUCT;
END_TYPE

TYPE "UDT1853_FLT_MeteringPump"
VERSION : 0.1
   STRUCT
      FLT_Prepressure : Bool;   // Fault prepressure metering pump too low (1)
      FLT_Motorprotection : Bool;   // Fault motorprotection metering pump (1)
      FLT_Max_pressure : Bool;   // Fault component pressure metering pump too high (1)
      FLT_SpP_Runtime : Bool;   // Fault prepressure from feed pump too low (1)
      FLT_F_converter : Bool;   // Fault frequency converter motor metering pump (1)
      FLT_Ventilation : Bool;   // Fault motorprotection ventilation dirve of drive pump(3)
      FLT_Min_Level : Bool;   // Fault min level day tank (3)
      FLT_Min_Pressure : Bool;   // Fault min Pressure before mixinghead opens (1)
      FLT_PreAlarmBearing : Bool;   // Fault pre alarm ball bearing
      FLT_Tolerance_high : Bool;   // Fault: Tolerance of flow exceeded (3)
      FLT_Tolerance_low : Bool;   // Fault: Tolerance of flow dropped (3)
      FLT_FlowSDATimeOut : Bool;   // Fault: Time out quick pressure build up (3)
      Mes_Min_temp : Bool;   // Message: Min temperature to start pump not reached
      Mes_StartUpDelayFU : Bool;   // Message: Start up delay FU (4)
      FLT_AlarmBearing : Bool;   // Fault: Alarm ball bearing
      FLT_FlowControlAtLimit : Bool;   // Fault: Flow controler at upper limit (3)
      Mes_PumpDeselected : Bool;   // Message: Pump is deselected for maintenance purposes
      Mes_PumpDeselectedInt : Bool;   // Message: Pump is deselected and runs in interval mode
      FLT_MotorFan : Bool;   // Fault: Motorprotection external fan of motor (2)
      FLT_DeselectedCompReqest : Bool;   // Fault: The component is deselected but needed for the next shot (1)
      FLT_FlowControlAtLOWLimit : Bool;   // Fault: Flow controler at lower limit (3)
      FLT_MaxLTripTray : Bool;   // Maximum level triptray (3)
      Spare2_6 : Bool;
      Spare2_7 : Bool;
      Spare3_0 : Bool;
      Spare3_1 : Bool;
      Spare3_2 : Bool;
      Spare3_3 : Bool;
      Spare3_4 : Bool;
      Spare3_5 : Bool;
      Spare3_6 : Bool;
      Spare3_7 : Bool;
   END_STRUCT;
END_TYPE

TYPE "UDT1860_FLT_ServE-Cyl"
VERSION : 0.1
   STRUCT
      TorqueUpperLimit : Bool;
      TorqueLowerLimit : Bool;
      Operable : Bool;
      FLT_MotorProtectionFU : Bool;
      spare_04 : Bool;
      spare_05 : Bool;
      spare_06 : Bool;
      spare_07 : Bool;
      spare_08 : Bool;
      spare_09 : Bool;
      spare_010 : Bool;
      spare_011 : Bool;
      spare_012 : Bool;
      spare_013 : Bool;
      spare_014 : Bool;
      spare_015 : Bool;
   END_STRUCT;
END_TYPE

TYPE "UDT1861_FLT_CylManager"
VERSION : 0.1
   STRUCT
      FirstEntry : Word;
   END_STRUCT;
END_TYPE

TYPE "UDT1862_FLT_Cylinder"
VERSION : 0.1
   STRUCT
      FLT_P_VentingHyd : Bool;   // Störung bei der Druckentlastung zur Entlüftung der Hydraulik nach dem Dosieren
      FLT_PMax_Component : Bool;   // Störung der maximale Komponentendruck wurde überschritten
      FLT_MotorprotectFeedp : Bool;   // Störung der Versorgung oder des Motorschutzes der Speisepumpe
      FLT_FeP_Runtime : Bool;   // Störung der Vordruck für den Zylinder wurde innerhalb 10 sec. nicht erreicht
      FLT_L_MinScavenger : Bool;   // Störung der Füllstand für die Spülmittelpumpe wurde unterschritten
      FLT_FeedpPrepressure : Bool;   // Störung der Vordruck der Komponente für den Zylinder ist nicht groß genug
      FLT_MaxPresHydraulic : Bool;   // Störung: Der maximale Hydraulikdruck für die Zylinderbewegung ist überschritten
      FLT_SealingMonitoring : Bool;   // Störung: Bei der Ansteuerung zum Füllen Packungs- Druck überschritten
      FLT_CylinderEmptyShot : Bool;   // Störung: Zylinder ist leer vor Schussende
      FLT_LimitSwitch : Bool;   // Störung: Endschalter Zylinder Komponente gestört
      Spare_1_2 : Bool;
      Spare_1_3 : Bool;
      Spare_1_4 : Bool;
      Spare_1_5 : Bool;
      Spare_1_6 : Bool;
      Spare_1_7 : Bool;
   END_STRUCT;
END_TYPE

TYPE "UDT1863_FLT_CylTandem"
VERSION : 0.1
   STRUCT
      FLT_TANDEM_PISTON_END : Bool;   // error: end of cylinder reached, changeover not completed
      FLT_TANDEM_GDA_TIMEOUT : Bool;   // error: timeout at pressure build-up
      FLT_TANDEM_PRESSURE_VA : Bool;   // error: unexpected pressure values at changeover
      FLT_TANDEM_NO_PISTON : Bool;   // error: Metering selected but no piston ready (because both are filling)
      FLT_TANDEM_RESERVED5 : Bool;   // Reserve
      FLT_MotorProtectionFU : Bool;   // Motor protection frequence converter tandem cylinder
      Spare_0_6 : Bool;
      Spare_0_7 : Bool;
      Spare_1_0 : Bool;
      Spare_1_1 : Bool;
      Spare_1_2 : Bool;
      Spare_1_3 : Bool;
      Spare_1_4 : Bool;
      Spare_1_5 : Bool;
      Spare_1_6 : Bool;
      Spare_1_7 : Bool;
   END_STRUCT;
END_TYPE

TYPE "UDT1871_FLT_CPiston"
VERSION : 0.1
   STRUCT
      Forward_to_slow : Bool;   // The motion of the cleanig piston to forward end position is too slow (1)
      Back_to_slow : Bool;   // The motion of the cleanig piston to backward end position is too slow (1)
      IPS_defect : Bool;   // Fault of inductive proximity switch at cleaning piston (1)
      Lost_IPS_position : Bool;   // Fault of inductive proximity switch at cleaning piston during foaming (1)
      Not_defind : Bool;   // Cleaning Piston not defined
      Spare_0_5 : Bool;
      Spare_0_6 : Bool;
      Spare_0_7 : Bool;
      Contr_upper_Limit : Bool;   // Controller cleaning piston at upper limit
      Contr_lower_Limit : Bool;   // Controller cleaning piston at lower limit
      Spare_1_2 : Bool;
      Never_reach_frontPos : Bool;   // Cleaning Piston never reaches front position
      Never_reach_backPos : Bool;   // Cleaning Piston never reaches end position
      Leaves_HomePos : Bool;   // Cleaning Piston leaves home position without activation
      Spare_1_6 : Bool;
      Spare_1_7 : Bool;
   END_STRUCT;
END_TYPE

TYPE "UDT1873_FLT_CPistonMQMX"
VERSION : 0.1
   STRUCT
      Stoer_LFZRKVor_MQ : Bool;
      Stoer_LFZRKZurueck_MQ : Bool;
      Stoer_LFZDrosselVor_MQ : Bool;
      Stoer_LFZDrossZurueck_MQ : Bool;
      Stoer_Dosierstellung_MQ : Bool;
      Stoer_Grundstellung_MQ : Bool;
      Stoer_Initiatoren_MQ : Bool;
      Stoer_LFZRK_MX : Bool;
      Stoer_LFZDrossel_MX : Bool;
      Stoer_LFZDosierkolben_MX : Bool;
      Stoer_Dosierstellung_MX : Bool;
      Res_STG1 : Bool;
      Res_STG2 : Bool;
      Res_STG3 : Bool;
      Res_STG4 : Bool;
      Spare_17 : Bool;
   END_STRUCT;
END_TYPE

DATA_BLOCK "InterfaceVisu"   // DB1
{ S7_Optimized_Access := 'FALSE' }
VERSION : 0.1
   VAR
      ScreenNo01 : Int := 0;
      ScreenNo02 : Int := 888;
      ScreenNo03 : Int := 0;
      ScreenNo04 : Int := 0;
      ScreenNo05 : Int := 0;
      InterfaceVisu05 : Word := 16#0000;
      InterfaceVisu06 : Word := 16#0000;
      InterfaceVisu07 : Word := 16#0000;
      InterfaceVisu08 : Word := 16#0000;
      InterfaceVisu09 : Word := 16#0000;
      InterfaceVisu10 : Word := 16#0000;
      InterfaceVisu11 : Word := 16#0000;
      InterfaceVisu12 : Word := 16#0000;
      InterfaceVisu13 : Word := 16#0000;
      InterfaceVisu14 : Word := 16#0000;
      InterfaceVisu15 : Word := 16#0000;
      InterfaceVisu16 : Word := 16#0000;
      InterfaceVisu17 : Word := 16#0000;
      InterfaceVisu18 : Word := 16#0000;
      InterfaceVisu19 : Word := 16#0000;
      InterfaceVisu20 : Word := 16#0000;
      InterfaceVisu21 : Word := 16#0000;
      InterfaceVisu22 : Word := 16#0000;
      InterfaceVisu23 : Word := 16#0000;
      InterfaceVisu24 : Word := 16#0000;
      InterfaceVisu25 : Word := 16#0000;
      InterfaceVisu26 : Word := 16#0000;
      InterfaceVisu27 : Word := 16#0000;
      InterfaceVisu28 : Word := 16#0000;
      InterfaceVisu29 : Word := 16#0000;
      InterfaceVisu30 : Word := 16#0000;
      InterfaceVisu31 : Word := 16#0000;
      InterfaceVisu32 : Word := 16#0000;
      InterfaceVisu33 : Word := 16#0000;
      InterfaceVisu34 : Word := 16#0000;
      InterfaceVisu35 : Word := 16#0000;
      InterfaceVisu36 : Word := 16#0000;
      InterfaceVisu37 : Word := 16#0000;
      InterfaceVisu38 : Word := 16#0000;
      InterfaceVisu39 : Word := 16#0000;
      InterfaceVisu40 : Word := 16#0000;
      InterfaceVisu41 : Word := 16#0000;
      InterfaceVisu42 : Word := 16#0000;
      InterfaceVisu43 : Word := 16#0000;
      InterfaceVisu44 : Word := 16#0000;
      InterfaceVisu45 : Word := 16#0000;
      InterfaceVisu46 : Word := 16#0000;
      InterfaceVisu47 : Word := 16#0000;
      InterfaceVisu48 : Word := 16#0000;
      InterfaceVisu49 : Word := 16#0000;
      ReadWriteDeviceNo : Int := 1;
      CopyDeviceNO : Int := 0;
      Read : Bool := FALSE;
      Write : Bool := FALSE;
      Copy : Bool := FALSE;
      Delete : Bool := FALSE;
      SetHDValue : Bool := FALSE;
      PopUp_MH_No : Bool := FALSE;
      HPValuesSet : Bool := FALSE;
      SpareByte : Byte := 16#00;
      NameComp : Array[1..8] of String[20];
      CompAtMixinghead : Array[1..8] of Bool;   // For visibility of the flow value
      ToolNo : Int := 0;
      LastPartShot : Bool;   // Maximum of part shots created in mould editor
      LastTool : Bool;   // Last tool selected in mould editor
      TestBit01 : Bool;
      TestBit2 : Bool;
      TestBit3 : Bool;
      TestBit4 : Bool;
      TestBit5 : Bool;
      TestBit6 : Bool;
      Input : Int := 0;
      "2PoinMovementComp" : Array[1..8] of Bool;   // For visibility of the flow value
      RefComponentComp : Array[1..8] of Bool;   // For visibility of the flow value
      RefComponent : Int := 1;
      MinFlow : Array[1..6] of Real;   // Minimum mass flow of pump [g/sec]
      MaxFlow : Array[1..6] of Real;   // Maximum mass flow of pump [g/sec]
      MaxTotalFlow : Array[0..8] of Real;
      MH_No_for_HPValues : Int;
      MaxShottime : Real;
      MinShottime : Real;
      AmountPartShots : Int;
      AmountTools : Int;
      AmountAlloactionAutomatic : Int;   // Amount of tools in allocation list in automatic
   END_VAR
BEGIN
   NameComp[1] := 'Poly';
   NameComp[2] := 'Iso';
   NameComp[3] := '   ';
   NameComp[4] := '   ';
   NameComp[5] := '   ';
   NameComp[6] := '   ';
   NameComp[7] := '';
   NameComp[8] := '';
   CompAtMixinghead[1] := TRUE;
   CompAtMixinghead[2] := TRUE;
   CompAtMixinghead[3] := FALSE;
   CompAtMixinghead[4] := FALSE;
   CompAtMixinghead[5] := FALSE;
   CompAtMixinghead[6] := FALSE;
   CompAtMixinghead[7] := FALSE;
   CompAtMixinghead[8] := FALSE;
   "2PoinMovementComp"[1] := FALSE;
   "2PoinMovementComp"[2] := FALSE;
   "2PoinMovementComp"[3] := FALSE;
   "2PoinMovementComp"[4] := FALSE;
   "2PoinMovementComp"[5] := FALSE;
   "2PoinMovementComp"[6] := FALSE;
   "2PoinMovementComp"[7] := FALSE;
   "2PoinMovementComp"[8] := FALSE;
   RefComponentComp[1] := FALSE;
   RefComponentComp[2] := FALSE;
   RefComponentComp[3] := FALSE;
   RefComponentComp[4] := FALSE;
   RefComponentComp[5] := FALSE;
   RefComponentComp[6] := FALSE;
   RefComponentComp[7] := FALSE;
   RefComponentComp[8] := FALSE;
   MaxFlow[1] := 667.0;
   MaxFlow[2] := 667.0;
   MaxFlow[3] := 0.0;
   MaxFlow[4] := 0.0;
   MaxFlow[5] := 0.0;
   MaxFlow[6] := 0.0;
   MinFlow[1] := 667.0;
   MinFlow[2] := 667.0;
   MinFlow[3] := 0.0;
   MinFlow[4] := 0.0;
   MinFlow[5] := 0.0;
   MinFlow[6] := 0.0;
END_DATA_BLOCK

DATA_BLOCK "DB905_GWK"   // DB2
{ S7_Optimized_Access := 'TRUE' }
VERSION : 0.1
   VAR
      teco_cs_cw_e : Array[0..2] of "PB_TecoCS(CW)e_SW-IW";   // Einfaches Protokoll teco cs cw
      State : Array[0..2] of "UDT_State_GWK";
   END_VAR
BEGIN
END_DATA_BLOCK

DATA_BLOCK "TP-Bereichszeiger"   // DB3
{ S7_Optimized_Access := 'FALSE' }
VERSION : 0.1
   VAR
      Koordinierungsbereich : Struct
         Intern_Byte_0 : Byte := 16#00;
         Anlaufbit : Bool := TRUE;
         Betriebsart_offline : Bool := FALSE;
         Lebensbit : Bool := FALSE;
         Intern_Bit_1_3 : Bool := FALSE;
         Intern_Bit_1_4 : Bool := FALSE;
         Intern_Bit_1_5 : Bool := FALSE;
         Intern_Bit_1_6 : Bool := FALSE;
         Intern_Bit_1_7 : Bool := FALSE;
      END_STRUCT;
      Auftragsfach : Struct
         Auftragsnummer : Int := 0;
         Parameter_01 : Word := 16#0000;
         Parameter_02 : Word := 16#0000;
         Parameter_03 : Word := 16#0000;
      END_STRUCT;
      Datenfach : Struct
         Rezepturnummer : Int := 0;
         Datensatznummer : Int := 0;
         Intern_Word_2 : Word := 16#0000;
         Status : Int := 0;
         Intern_Word_4 : Word := 16#0000;
      END_STRUCT;
      Picturenumber : Struct
         Bildtyp : Word := 16#0001;
         Bildnummer : Int := 16#0018;
         Intern_Word_2 : Word := 16#0000;
         Eingabefeldnummer : Word := 16#0001;
         Intern_Word_4 : Word := 16#0000;
      END_STRUCT;
      Date_Time : Struct
         Start_AG_Transfer : Bool := FALSE;
         Reserve_1 : Bool := FALSE;
         Reserve_2 : Bool := FALSE;
         Reserve_3 : Bool := FALSE;
         Reserve_4 : Bool := FALSE;
         Reserve_5 : Bool := FALSE;
         Reserve_6 : Bool := FALSE;
         Reserve_7 : Bool := FALSE;
         SetTime : DTL := DTL#1970-01-01-00:00:00;
         ActTime : DTL := DTL#2016-12-19-10:16:07.659621044;
         reserviert : DWord := 16#0000_0000;
      END_STRUCT;
   END_VAR
BEGIN
END_DATA_BLOCK

DATA_BLOCK "DB1009_TT_Config"   // DB4
{ S7_Optimized_Access := 'FALSE' }
VERSION : 0.1
   VAR
      Bit : Struct
         WithTT : Bool := TRUE;
         WithRobot : Bool := FALSE;
      END_STRUCT;
      AmountOfSegment : Int := 6;
   END_VAR
BEGIN
END_DATA_BLOCK

DATA_BLOCK "DB005_RS<->Extern"   // DB5
TITLE = Interface signals between PU and external plant
{ S7_Optimized_Access := 'FALSE' }
AUTHOR : KT242